   11: [NEQ(MV_MV12R.DriveBits,0) OTE(MV_MV12R.CW.[CWD.AUTODRV]) ,[XIC(MV_MV12R.CW.[CWD.AUTODRV]) XIO(MV_MV12R.CW.[CWD.MANUAL]) ,XIC(MV_MV12R.CW.[CWD.MANDRV]) XIC(MV_MV12R.CW.[CWD.MANUAL]) ] OTE(MV_MV12R.CW.[CWD.OUTPUT]) ,XIC(MV_MV12R.CW.[CWD.OUTPUT]) OTE(MV_MV12R_D) ,XIC(S:FS) [OTU(MV_MV12R.CW.[CWD.MANUAL]) ,LEQ(MV_MV12R.CheckTime,0) MOV(Default_Check_Time,MV_MV12R.CheckTime) ] ,[[XIC(MV_MV12R_R) XIO(Item_Simulation_Flag) ,XIC(Item_Simulation_Flag) [XIC(MV_MV12R.CW.[CWD.OUTPUT]) XIO(MV_MV12R.CW.[CWD.SIMFAIL]) ,XIO(MV_MV12R.CW.[CWD.OUTPUT]) XIC(MV_MV12R.CW.[CWD.SIMFAIL]) ] ] OTE(MV_MV12R.CW.[CWD.RUNFB]) ,[XIC(Item_Simulation_Flag) ,XIC(MV_MV12R.CW.[CWD.CHECKOFF]) ,XIC(Unused_Healthy_Feedback) ] OTE(MV_MV12R.CW.[CWD.HEALTHYFB]) ,[XIC(Item_Simulation_Flag) ,XIC(MV_MV12R.CW.[CWD.CHECKOFF]) ,XIC(Unused_NotTripped_Feedback) ] OTE(MV_MV12R.CW.[CWD.NOTTRIPPEDFB]) ] ,[XIC(MV_MV12R.CW.[CWD.AUTODRV]) XIO(MV_MV12R.CW.[CWD.PREVSCAN]) ,XIO(MV_MV12R.CW.[CWD.AUTODRV]) XIC(MV_MV12R.CW.[CWD.PREVSCAN]) ] CLR(MV_MV12R.CheckTimer) ,XIC(One_Second_One_Scan) LES(MV_MV12R.CheckTimer,MV_MV12R.CheckTime) ADD(MV_MV12R.CheckTimer,1,MV_MV12R.CheckTimer) ,XIO(MV_MV12R.CW.[CWD.FAULT]) OTU(MV_MV12R.CW.[CWD.FAULTLOGGED]) ,[GEQ(MV_MV12R.CheckTimer,MV_MV12R.CheckTime) [XIC(MV_MV12R.CW.[CWD.OUTPUT]) XIO(MV_MV12R.CW.[CWD.RUNFB]) ,XIO(MV_MV12R.CW.[CWD.OUTPUT]) XIC(MV_MV12R.CW.[CWD.RUNFB]) ] ,XIO(MV_MV12R.CW.[CWD.HEALTHYFB]) ,XIO(MV_MV12R.CW.[CWD.NOTTRIPPEDFB]) ,XIC(MV_MV12R.CW.[CWD.FAULT]) XIC(Item_Faults_Are_Latched) ,XIC(MV_MV12R.CW.[CWD.HIGHLIGHT]) ] XIO(MV_MV12R.CW.[CWD.CHECKOFF]) XIO(Alarm_Reset) [OTE(MV_MV12R.CW.[CWD.FAULT]) ,ALMD(MV_MV12R_ALARM,0,0,0,0) ] ,XIC(MV_MV12R.CW.[CWD.OUTPUT]) OTE(MV_MV12R.CW.[CWD.PREVSCAN]) ,XIC(MV_MV12R.CW.[CWD.FAULT]) EQU(Scada_Pump_Fault_No,0) XIO(MV_MV12R.CW.[CWD.FAULTLOGGED]) [MOV(20001,Scada_Pump_Fault_No) ,OTL(MV_MV12R.CW.[CWD.FAULTLOGGED]) ] ,XIO(MV_MV12R.CW.[CWD.HEALTHYFB]) EQU(Scada_Pump_H_Fault_No,0) XIO(MV_MV12R.CW.[CWD.HEALTHYFAULTLOGGED]) [MOV(20001,Scada_Pump_H_Fault_No) ,OTL(MV_MV12R.CW.[CWD.HEALTHYFAULTLOGGED]) ] ,XIO(MV_MV12R.CW.[CWD.NOTTRIPPEDFB]) EQU(Scada_Pump_H_Fault_No,0) XIO(MV_MV12R.CW.[CWD.TRIPPEDFAULTLOGGED]) [MOV(20001,Scada_Pump_T_Fault_No) ,OTL(MV_MV12R.CW.[CWD.TRIPPEDFAULTLOGGED]) ] ];
   12: [NEQ(MV_MV13R.DriveBits,0) OTE(MV_MV13R.CW.[CWD.AUTODRV]) ,[XIC(MV_MV13R.CW.[CWD.AUTODRV]) XIO(MV_MV13R.CW.[CWD.MANUAL]) ,XIC(MV_MV13R.CW.[CWD.MANDRV]) XIC(MV_MV13R.CW.[CWD.MANUAL]) ] OTE(MV_MV13R.CW.[CWD.OUTPUT]) ,XIC(MV_MV13R.CW.[CWD.OUTPUT]) OTE(MV_MV13R_D) ,XIC(S:FS) [OTU(MV_MV13R.CW.[CWD.MANUAL]) ,LEQ(MV_MV13R.CheckTime,0) MOV(Default_Check_Time,MV_MV13R.CheckTime) ] ,[[XIC(MV_MV13R_R) XIO(Item_Simulation_Flag) ,XIC(Item_Simulation_Flag) [XIC(MV_MV13R.CW.[CWD.OUTPUT]) XIO(MV_MV13R.CW.[CWD.SIMFAIL]) ,XIO(MV_MV13R.CW.[CWD.OUTPUT]) XIC(MV_MV13R.CW.[CWD.SIMFAIL]) ] ] OTE(MV_MV13R.CW.[CWD.RUNFB]) ,[XIC(Item_Simulation_Flag) ,XIC(MV_MV13R.CW.[CWD.CHECKOFF]) ,XIC(Unused_Healthy_Feedback) ] OTE(MV_MV13R.CW.[CWD.HEALTHYFB]) ,[XIC(Item_Simulation_Flag) ,XIC(MV_MV13R.CW.[CWD.CHECKOFF]) ,XIC(Unused_NotTripped_Feedback) ] OTE(MV_MV13R.CW.[CWD.NOTTRIPPEDFB]) ] ,[XIC(MV_MV13R.CW.[CWD.AUTODRV]) XIO(MV_MV13R.CW.[CWD.PREVSCAN]) ,XIO(MV_MV13R.CW.[CWD.AUTODRV]) XIC(MV_MV13R.CW.[CWD.PREVSCAN]) ] CLR(MV_MV13R.CheckTimer) ,XIC(One_Second_One_Scan) LES(MV_MV13R.CheckTimer,MV_MV13R.CheckTime) ADD(MV_MV13R.CheckTimer,1,MV_MV13R.CheckTimer) ,XIO(MV_MV13R.CW.[CWD.FAULT]) OTU(MV_MV13R.CW.[CWD.FAULTLOGGED]) ,[GEQ(MV_MV13R.CheckTimer,MV_MV13R.CheckTime) [XIC(MV_MV13R.CW.[CWD.OUTPUT]) XIO(MV_MV13R.CW.[CWD.RUNFB]) ,XIO(MV_MV13R.CW.[CWD.OUTPUT]) XIC(MV_MV13R.CW.[CWD.RUNFB]) ] ,XIO(MV_MV13R.CW.[CWD.HEALTHYFB]) ,XIO(MV_MV13R.CW.[CWD.NOTTRIPPEDFB]) ,XIC(MV_MV13R.CW.[CWD.FAULT]) XIC(Item_Faults_Are_Latched) ,XIC(MV_MV13R.CW.[CWD.HIGHLIGHT]) ] XIO(MV_MV13R.CW.[CWD.CHECKOFF]) XIO(Alarm_Reset) [OTE(MV_MV13R.CW.[CWD.FAULT]) ,ALMD(MV_MV13R_ALARM,0,0,0,0) ] ,XIC(MV_MV13R.CW.[CWD.OUTPUT]) OTE(MV_MV13R.CW.[CWD.PREVSCAN]) ,XIC(MV_MV13R.CW.[CWD.FAULT]) EQU(Scada_Pump_Fault_No,0) XIO(MV_MV13R.CW.[CWD.FAULTLOGGED]) [MOV(20001,Scada_Pump_Fault_No) ,OTL(MV_MV13R.CW.[CWD.FAULTLOGGED]) ] ,XIO(MV_MV13R.CW.[CWD.HEALTHYFB]) EQU(Scada_Pump_H_Fault_No,0) XIO(MV_MV13R.CW.[CWD.HEALTHYFAULTLOGGED]) [MOV(20001,Scada_Pump_H_Fault_No) ,OTL(MV_MV13R.CW.[CWD.HEALTHYFAULTLOGGED]) ] ,XIO(MV_MV13R.CW.[CWD.NOTTRIPPEDFB]) EQU(Scada_Pump_H_Fault_No,0) XIO(MV_MV13R.CW.[CWD.TRIPPEDFAULTLOGGED]) [MOV(20001,Scada_Pump_T_Fault_No) ,OTL(MV_MV13R.CW.[CWD.TRIPPEDFAULTLOGGED]) ] ];
   13: [NEQ(MV_MV14R.DriveBits,0) OTE(MV_MV14R.CW.[CWD.AUTODRV]) ,[XIC(MV_MV14R.CW.[CWD.AUTODRV]) XIO(MV_MV14R.CW.[CWD.MANUAL]) ,XIC(MV_MV14R.CW.[CWD.MANDRV]) XIC(MV_MV14R.CW.[CWD.MANUAL]) ] OTE(MV_MV14R.CW.[CWD.OUTPUT]) ,XIC(MV_MV14R.CW.[CWD.OUTPUT]) OTE(MV_MV14R_D) ,XIC(S:FS) [OTU(MV_MV14R.CW.[CWD.MANUAL]) ,LEQ(MV_MV14R.CheckTime,0) MOV(Default_Check_Time,MV_MV14R.CheckTime) ] ,[[XIC(MV_MV14R_R) XIO(Item_Simulation_Flag) ,XIC(Item_Simulation_Flag) [XIC(MV_MV14R.CW.[CWD.OUTPUT]) XIO(MV_MV14R.CW.[CWD.SIMFAIL]) ,XIO(MV_MV14R.CW.[CWD.OUTPUT]) XIC(MV_MV14R.CW.[CWD.SIMFAIL]) ] ] OTE(MV_MV14R.CW.[CWD.RUNFB]) ,[XIC(Item_Simulation_Flag) ,XIC(MV_MV14R.CW.[CWD.CHECKOFF]) ,XIC(Unused_Healthy_Feedback) ] OTE(MV_MV14R.CW.[CWD.HEALTHYFB]) ,[XIC(Item_Simulation_Flag) ,XIC(MV_MV14R.CW.[CWD.CHECKOFF]) ,XIC(Unused_NotTripped_Feedback) ] OTE(MV_MV14R.CW.[CWD.NOTTRIPPEDFB]) ] ,[XIC(MV_MV14R.CW.[CWD.AUTODRV]) XIO(MV_MV14R.CW.[CWD.PREVSCAN]) ,XIO(MV_MV14R.CW.[CWD.AUTODRV]) XIC(MV_MV14R.CW.[CWD.PREVSCAN]) ] CLR(MV_MV14R.CheckTimer) ,XIC(One_Second_One_Scan) LES(MV_MV14R.CheckTimer,MV_MV14R.CheckTime) ADD(MV_MV14R.CheckTimer,1,MV_MV14R.CheckTimer) ,XIO(MV_MV14R.CW.[CWD.FAULT]) OTU(MV_MV14R.CW.[CWD.FAULTLOGGED]) ,[GEQ(MV_MV14R.CheckTimer,MV_MV14R.CheckTime) [XIC(MV_MV14R.CW.[CWD.OUTPUT]) XIO(MV_MV14R.CW.[CWD.RUNFB]) ,XIO(MV_MV14R.CW.[CWD.OUTPUT]) XIC(MV_MV14R.CW.[CWD.RUNFB]) ] ,XIO(MV_MV14R.CW.[CWD.HEALTHYFB]) ,XIO(MV_MV14R.CW.[CWD.NOTTRIPPEDFB]) ,XIC(MV_MV14R.CW.[CWD.FAULT]) XIC(Item_Faults_Are_Latched) ,XIC(MV_MV14R.CW.[CWD.HIGHLIGHT]) ] XIO(MV_MV14R.CW.[CWD.CHECKOFF]) XIO(Alarm_Reset) [OTE(MV_MV14R.CW.[CWD.FAULT]) ,ALMD(MV_MV14R_ALARM,0,0,0,0) ] ,XIC(MV_MV14R.CW.[CWD.OUTPUT]) OTE(MV_MV14R.CW.[CWD.PREVSCAN]) ,XIC(MV_MV14R.CW.[CWD.FAULT]) EQU(Scada_Pump_Fault_No,0) XIO(MV_MV14R.CW.[CWD.FAULTLOGGED]) [MOV(20001,Scada_Pump_Fault_No) ,OTL(MV_MV14R.CW.[CWD.FAULTLOGGED]) ] ,XIO(MV_MV14R.CW.[CWD.HEALTHYFB]) EQU(Scada_Pump_H_Fault_No,0) XIO(MV_MV14R.CW.[CWD.HEALTHYFAULTLOGGED]) [MOV(20001,Scada_Pump_H_Fault_No) ,OTL(MV_MV14R.CW.[CWD.HEALTHYFAULTLOGGED]) ] ,XIO(MV_MV14R.CW.[CWD.NOTTRIPPEDFB]) EQU(Scada_Pump_H_Fault_No,0) XIO(MV_MV14R.CW.[CWD.TRIPPEDFAULTLOGGED]) [MOV(20001,Scada_Pump_T_Fault_No) ,OTL(MV_MV14R.CW.[CWD.TRIPPEDFAULTLOGGED]) ] ];
   14: [NEQ(MV_MV15R.DriveBits,0) OTE(MV_MV15R.CW.[CWD.AUTODRV]) ,[XIC(MV_MV15R.CW.[CWD.AUTODRV]) XIO(MV_MV15R.CW.[CWD.MANUAL]) ,XIC(MV_MV15R.CW.[CWD.MANDRV]) XIC(MV_MV15R.CW.[CWD.MANUAL]) ] OTE(MV_MV15R.CW.[CWD.OUTPUT]) ,XIC(MV_MV15R.CW.[CWD.OUTPUT]) OTE(MV_MV15R_D) ,XIC(S:FS) [OTU(MV_MV15R.CW.[CWD.MANUAL]) ,LEQ(MV_MV15R.CheckTime,0) MOV(Default_Check_Time,MV_MV15R.CheckTime) ] ,[[XIC(MV_MV15R_R) XIO(Item_Simulation_Flag) ,XIC(Item_Simulation_Flag) [XIC(MV_MV15R.CW.[CWD.OUTPUT]) XIO(MV_MV15R.CW.[CWD.SIMFAIL]) ,XIO(MV_MV15R.CW.[CWD.OUTPUT]) XIC(MV_MV15R.CW.[CWD.SIMFAIL]) ] ] OTE(MV_MV15R.CW.[CWD.RUNFB]) ,[XIC(Item_Simulation_Flag) ,XIC(MV_MV15R.CW.[CWD.CHECKOFF]) ,XIC(Unused_Healthy_Feedback) ] OTE(MV_MV15R.CW.[CWD.HEALTHYFB]) ,[XIC(Item_Simulation_Flag) ,XIC(MV_MV15R.CW.[CWD.CHECKOFF]) ,XIC(Unused_NotTripped_Feedback) ] OTE(MV_MV15R.CW.[CWD.NOTTRIPPEDFB]) ] ,[XIC(MV_MV15R.CW.[CWD.AUTODRV]) XIO(MV_MV15R.CW.[CWD.PREVSCAN]) ,XIO(MV_MV15R.CW.[CWD.AUTODRV]) XIC(MV_MV15R.CW.[CWD.PREVSCAN]) ] CLR(MV_MV15R.CheckTimer) ,XIC(One_Second_One_Scan) LES(MV_MV15R.CheckTimer,MV_MV15R.CheckTime) ADD(MV_MV15R.CheckTimer,1,MV_MV15R.CheckTimer) ,XIO(MV_MV15R.CW.[CWD.FAULT]) OTU(MV_MV15R.CW.[CWD.FAULTLOGGED]) ,[GEQ(MV_MV15R.CheckTimer,MV_MV15R.CheckTime) [XIC(MV_MV15R.CW.[CWD.OUTPUT]) XIO(MV_MV15R.CW.[CWD.RUNFB]) ,XIO(MV_MV15R.CW.[CWD.OUTPUT]) XIC(MV_MV15R.CW.[CWD.RUNFB]) ] ,XIO(MV_MV15R.CW.[CWD.HEALTHYFB]) ,XIO(MV_MV15R.CW.[CWD.NOTTRIPPEDFB]) ,XIC(MV_MV15R.CW.[CWD.FAULT]) XIC(Item_Faults_Are_Latched) ,XIC(MV_MV15R.CW.[CWD.HIGHLIGHT]) ] XIO(MV_MV15R.CW.[CWD.CHECKOFF]) XIO(Alarm_Reset) [OTE(MV_MV15R.CW.[CWD.FAULT]) ,ALMD(MV_MV15R_ALARM,0,0,0,0) ] ,XIC(MV_MV15R.CW.[CWD.OUTPUT]) OTE(MV_MV15R.CW.[CWD.PREVSCAN]) ,XIC(MV_MV15R.CW.[CWD.FAULT]) EQU(Scada_Pump_Fault_No,0) XIO(MV_MV15R.CW.[CWD.FAULTLOGGED]) [MOV(20001,Scada_Pump_Fault_No) ,OTL(MV_MV15R.CW.[CWD.FAULTLOGGED]) ] ,XIO(MV_MV15R.CW.[CWD.HEALTHYFB]) EQU(Scada_Pump_H_Fault_No,0) XIO(MV_MV15R.CW.[CWD.HEALTHYFAULTLOGGED]) [MOV(20001,Scada_Pump_H_Fault_No) ,OTL(MV_MV15R.CW.[CWD.HEALTHYFAULTLOGGED]) ] ,XIO(MV_MV15R.CW.[CWD.NOTTRIPPEDFB]) EQU(Scada_Pump_H_Fault_No,0) XIO(MV_MV15R.CW.[CWD.TRIPPEDFAULTLOGGED]) [MOV(20001,Scada_Pump_T_Fault_No) ,OTL(MV_MV15R.CW.[CWD.TRIPPEDFAULTLOGGED]) ] ];
   15: [NEQ(MV_MV16R.DriveBits,0) OTE(MV_MV16R.CW.[CWD.AUTODRV]) ,[XIC(MV_MV16R.CW.[CWD.AUTODRV]) XIO(MV_MV16R.CW.[CWD.MANUAL]) ,XIC(MV_MV16R.CW.[CWD.MANDRV]) XIC(MV_MV16R.CW.[CWD.MANUAL]) ] OTE(MV_MV16R.CW.[CWD.OUTPUT]) ,XIC(MV_MV16R.CW.[CWD.OUTPUT]) OTE(MV_MV16R_D) ,XIC(S:FS) [OTU(MV_MV16R.CW.[CWD.MANUAL]) ,LEQ(MV_MV16R.CheckTime,0) MOV(Default_Check_Time,MV_MV16R.CheckTime) ] ,[[XIC(MV_MV16R_R) XIO(Item_Simulation_Flag) ,XIC(Item_Simulation_Flag) [XIC(MV_MV16R.CW.[CWD.OUTPUT]) XIO(MV_MV16R.CW.[CWD.SIMFAIL]) ,XIO(MV_MV16R.CW.[CWD.OUTPUT]) XIC(MV_MV16R.CW.[CWD.SIMFAIL]) ] ] OTE(MV_MV16R.CW.[CWD.RUNFB]) ,[XIC(Item_Simulation_Flag) ,XIC(MV_MV16R.CW.[CWD.CHECKOFF]) ,XIC(Unused_Healthy_Feedback) ] OTE(MV_MV16R.CW.[CWD.HEALTHYFB]) ,[XIC(Item_Simulation_Flag) ,XIC(MV_MV16R.CW.[CWD.CHECKOFF]) ,XIC(Unused_NotTripped_Feedback) ] OTE(MV_MV16R.CW.[CWD.NOTTRIPPEDFB]) ] ,[XIC(MV_MV16R.CW.[CWD.AUTODRV]) XIO(MV_MV16R.CW.[CWD.PREVSCAN]) ,XIO(MV_MV16R.CW.[CWD.AUTODRV]) XIC(MV_MV16R.CW.[CWD.PREVSCAN]) ] CLR(MV_MV16R.CheckTimer) ,XIC(One_Second_One_Scan) LES(MV_MV16R.CheckTimer,MV_MV16R.CheckTime) ADD(MV_MV16R.CheckTimer,1,MV_MV16R.CheckTimer) ,XIO(MV_MV16R.CW.[CWD.FAULT]) OTU(MV_MV16R.CW.[CWD.FAULTLOGGED]) ,[GEQ(MV_MV16R.CheckTimer,MV_MV16R.CheckTime) [XIC(MV_MV16R.CW.[CWD.OUTPUT]) XIO(MV_MV16R.CW.[CWD.RUNFB]) ,XIO(MV_MV16R.CW.[CWD.OUTPUT]) XIC(MV_MV16R.CW.[CWD.RUNFB]) ] ,XIO(MV_MV16R.CW.[CWD.HEALTHYFB]) ,XIO(MV_MV16R.CW.[CWD.NOTTRIPPEDFB]) ,XIC(MV_MV16R.CW.[CWD.FAULT]) XIC(Item_Faults_Are_Latched) ,XIC(MV_MV16R.CW.[CWD.HIGHLIGHT]) ] XIO(MV_MV16R.CW.[CWD.CHECKOFF]) XIO(Alarm_Reset) [OTE(MV_MV16R.CW.[CWD.FAULT]) ,ALMD(MV_MV16R_ALARM,0,0,0,0) ] ,XIC(MV_MV16R.CW.[CWD.OUTPUT]) OTE(MV_MV16R.CW.[CWD.PREVSCAN]) ,XIC(MV_MV16R.CW.[CWD.FAULT]) EQU(Scada_Pump_Fault_No,0) XIO(MV_MV16R.CW.[CWD.FAULTLOGGED]) [MOV(20001,Scada_Pump_Fault_No) ,OTL(MV_MV16R.CW.[CWD.FAULTLOGGED]) ] ,XIO(MV_MV16R.CW.[CWD.HEALTHYFB]) EQU(Scada_Pump_H_Fault_No,0) XIO(MV_MV16R.CW.[CWD.HEALTHYFAULTLOGGED]) [MOV(20001,Scada_Pump_H_Fault_No) ,OTL(MV_MV16R.CW.[CWD.HEALTHYFAULTLOGGED]) ] ,XIO(MV_MV16R.CW.[CWD.NOTTRIPPEDFB]) EQU(Scada_Pump_H_Fault_No,0) XIO(MV_MV16R.CW.[CWD.TRIPPEDFAULTLOGGED]) [MOV(20001,Scada_Pump_T_Fault_No) ,OTL(MV_MV16R.CW.[CWD.TRIPPEDFAULTLOGGED]) ] ];
   16: [NEQ(MV_MV17R.DriveBits,0) OTE(MV_MV17R.CW.[CWD.AUTODRV]) ,[XIC(MV_MV17R.CW.[CWD.AUTODRV]) XIO(MV_MV17R.CW.[CWD.MANUAL]) ,XIC(MV_MV17R.CW.[CWD.MANDRV]) XIC(MV_MV17R.CW.[CWD.MANUAL]) ] OTE(MV_MV17R.CW.[CWD.OUTPUT]) ,XIC(MV_MV17R.CW.[CWD.OUTPUT]) OTE(MV_MV17R_D) ,XIC(S:FS) [OTU(MV_MV17R.CW.[CWD.MANUAL]) ,LEQ(MV_MV17R.CheckTime,0) MOV(Default_Check_Time,MV_MV17R.CheckTime) ] ,[[XIC(MV_MV17R_R) XIO(Item_Simulation_Flag) ,XIC(Item_Simulation_Flag) [XIC(MV_MV17R.CW.[CWD.OUTPUT]) XIO(MV_MV17R.CW.[CWD.SIMFAIL]) ,XIO(MV_MV17R.CW.[CWD.OUTPUT]) XIC(MV_MV17R.CW.[CWD.SIMFAIL]) ] ] OTE(MV_MV17R.CW.[CWD.RUNFB]) ,[XIC(Item_Simulation_Flag) ,XIC(MV_MV17R.CW.[CWD.CHECKOFF]) ,XIC(Unused_Healthy_Feedback) ] OTE(MV_MV17R.CW.[CWD.HEALTHYFB]) ,[XIC(Item_Simulation_Flag) ,XIC(MV_MV17R.CW.[CWD.CHECKOFF]) ,XIC(Unused_NotTripped_Feedback) ] OTE(MV_MV17R.CW.[CWD.NOTTRIPPEDFB]) ] ,[XIC(MV_MV17R.CW.[CWD.AUTODRV]) XIO(MV_MV17R.CW.[CWD.PREVSCAN]) ,XIO(MV_MV17R.CW.[CWD.AUTODRV]) XIC(MV_MV17R.CW.[CWD.PREVSCAN]) ] CLR(MV_MV17R.CheckTimer) ,XIC(One_Second_One_Scan) LES(MV_MV17R.CheckTimer,MV_MV17R.CheckTime) ADD(MV_MV17R.CheckTimer,1,MV_MV17R.CheckTimer) ,XIO(MV_MV17R.CW.[CWD.FAULT]) OTU(MV_MV17R.CW.[CWD.FAULTLOGGED]) ,[GEQ(MV_MV17R.CheckTimer,MV_MV17R.CheckTime) [XIC(MV_MV17R.CW.[CWD.OUTPUT]) XIO(MV_MV17R.CW.[CWD.RUNFB]) ,XIO(MV_MV17R.CW.[CWD.OUTPUT]) XIC(MV_MV17R.CW.[CWD.RUNFB]) ] ,XIO(MV_MV17R.CW.[CWD.HEALTHYFB]) ,XIO(MV_MV17R.CW.[CWD.NOTTRIPPEDFB]) ,XIC(MV_MV17R.CW.[CWD.FAULT]) XIC(Item_Faults_Are_Latched) ,XIC(MV_MV17R.CW.[CWD.HIGHLIGHT]) ] XIO(MV_MV17R.CW.[CWD.CHECKOFF]) XIO(Alarm_Reset) [OTE(MV_MV17R.CW.[CWD.FAULT]) ,ALMD(MV_MV17R_ALARM,0,0,0,0) ] ,XIC(MV_MV17R.CW.[CWD.OUTPUT]) OTE(MV_MV17R.CW.[CWD.PREVSCAN]) ,XIC(MV_MV17R.CW.[CWD.FAULT]) EQU(Scada_Pump_Fault_No,0) XIO(MV_MV17R.CW.[CWD.FAULTLOGGED]) [MOV(20001,Scada_Pump_Fault_No) ,OTL(MV_MV17R.CW.[CWD.FAULTLOGGED]) ] ,XIO(MV_MV17R.CW.[CWD.HEALTHYFB]) EQU(Scada_Pump_H_Fault_No,0) XIO(MV_MV17R.CW.[CWD.HEALTHYFAULTLOGGED]) [MOV(20001,Scada_Pump_H_Fault_No) ,OTL(MV_MV17R.CW.[CWD.HEALTHYFAULTLOGGED]) ] ,XIO(MV_MV17R.CW.[CWD.NOTTRIPPEDFB]) EQU(Scada_Pump_H_Fault_No,0) XIO(MV_MV17R.CW.[CWD.TRIPPEDFAULTLOGGED]) [MOV(20001,Scada_Pump_T_Fault_No) ,OTL(MV_MV17R.CW.[CWD.TRIPPEDFAULTLOGGED]) ] ];
   17: [NEQ(MV_MV18R.DriveBits,0) OTE(MV_MV18R.CW.[CWD.AUTODRV]) ,[XIC(MV_MV18R.CW.[CWD.AUTODRV]) XIO(MV_MV18R.CW.[CWD.MANUAL]) ,XIC(MV_MV18R.CW.[CWD.MANDRV]) XIC(MV_MV18R.CW.[CWD.MANUAL]) ] OTE(MV_MV18R.CW.[CWD.OUTPUT]) ,XIC(MV_MV18R.CW.[CWD.OUTPUT]) OTE(MV_MV18R_D) ,XIC(S:FS) [OTU(MV_MV18R.CW.[CWD.MANUAL]) ,LEQ(MV_MV18R.CheckTime,0) MOV(Default_Check_Time,MV_MV18R.CheckTime) ] ,[[XIC(MV_MV18R_R) XIO(Item_Simulation_Flag) ,XIC(Item_Simulation_Flag) [XIC(MV_MV18R.CW.[CWD.OUTPUT]) XIO(MV_MV18R.CW.[CWD.SIMFAIL]) ,XIO(MV_MV18R.CW.[CWD.OUTPUT]) XIC(MV_MV18R.CW.[CWD.SIMFAIL]) ] ] OTE(MV_MV18R.CW.[CWD.RUNFB]) ,[XIC(Item_Simulation_Flag) ,XIC(MV_MV18R.CW.[CWD.CHECKOFF]) ,XIC(Unused_Healthy_Feedback) ] OTE(MV_MV18R.CW.[CWD.HEALTHYFB]) ,[XIC(Item_Simulation_Flag) ,XIC(MV_MV18R.CW.[CWD.CHECKOFF]) ,XIC(Unused_NotTripped_Feedback) ] OTE(MV_MV18R.CW.[CWD.NOTTRIPPEDFB]) ] ,[XIC(MV_MV18R.CW.[CWD.AUTODRV]) XIO(MV_MV18R.CW.[CWD.PREVSCAN]) ,XIO(MV_MV18R.CW.[CWD.AUTODRV]) XIC(MV_MV18R.CW.[CWD.PREVSCAN]) ] CLR(MV_MV18R.CheckTimer) ,XIC(One_Second_One_Scan) LES(MV_MV18R.CheckTimer,MV_MV18R.CheckTime) ADD(MV_MV18R.CheckTimer,1,MV_MV18R.CheckTimer) ,XIO(MV_MV18R.CW.[CWD.FAULT]) OTU(MV_MV18R.CW.[CWD.FAULTLOGGED]) ,[GEQ(MV_MV18R.CheckTimer,MV_MV18R.CheckTime) [XIC(MV_MV18R.CW.[CWD.OUTPUT]) XIO(MV_MV18R.CW.[CWD.RUNFB]) ,XIO(MV_MV18R.CW.[CWD.OUTPUT]) XIC(MV_MV18R.CW.[CWD.RUNFB]) ] ,XIO(MV_MV18R.CW.[CWD.HEALTHYFB]) ,XIO(MV_MV18R.CW.[CWD.NOTTRIPPEDFB]) ,XIC(MV_MV18R.CW.[CWD.FAULT]) XIC(Item_Faults_Are_Latched) ,XIC(MV_MV18R.CW.[CWD.HIGHLIGHT]) ] XIO(MV_MV18R.CW.[CWD.CHECKOFF]) XIO(Alarm_Reset) [OTE(MV_MV18R.CW.[CWD.FAULT]) ,ALMD(MV_MV18R_ALARM,0,0,0,0) ] ,XIC(MV_MV18R.CW.[CWD.OUTPUT]) OTE(MV_MV18R.CW.[CWD.PREVSCAN]) ,XIC(MV_MV18R.CW.[CWD.FAULT]) EQU(Scada_Pump_Fault_No,0) XIO(MV_MV18R.CW.[CWD.FAULTLOGGED]) [MOV(20001,Scada_Pump_Fault_No) ,OTL(MV_MV18R.CW.[CWD.FAULTLOGGED]) ] ,XIO(MV_MV18R.CW.[CWD.HEALTHYFB]) EQU(Scada_Pump_H_Fault_No,0) XIO(MV_MV18R.CW.[CWD.HEALTHYFAULTLOGGED]) [MOV(20001,Scada_Pump_H_Fault_No) ,OTL(MV_MV18R.CW.[CWD.HEALTHYFAULTLOGGED]) ] ,XIO(MV_MV18R.CW.[CWD.NOTTRIPPEDFB]) EQU(Scada_Pump_H_Fault_No,0) XIO(MV_MV18R.CW.[CWD.TRIPPEDFAULTLOGGED]) [MOV(20001,Scada_Pump_T_Fault_No) ,OTL(MV_MV18R.CW.[CWD.TRIPPEDFAULTLOGGED]) ] ];
   18: [NEQ(MV_MV19R.DriveBits,0) OTE(MV_MV19R.CW.[CWD.AUTODRV]) ,[XIC(MV_MV19R.CW.[CWD.AUTODRV]) XIO(MV_MV19R.CW.[CWD.MANUAL]) ,XIC(MV_MV19R.CW.[CWD.MANDRV]) XIC(MV_MV19R.CW.[CWD.MANUAL]) ] OTE(MV_MV19R.CW.[CWD.OUTPUT]) ,XIC(MV_MV19R.CW.[CWD.OUTPUT]) OTE(MV_MV19R_D) ,XIC(S:FS) [OTU(MV_MV19R.CW.[CWD.MANUAL]) ,LEQ(MV_MV19R.CheckTime,0) MOV(Default_Check_Time,MV_MV19R.CheckTime) ] ,[[XIC(MV_MV19R_R) XIO(Item_Simulation_Flag) ,XIC(Item_Simulation_Flag) [XIC(MV_MV19R.CW.[CWD.OUTPUT]) XIO(MV_MV19R.CW.[CWD.SIMFAIL]) ,XIO(MV_MV19R.CW.[CWD.OUTPUT]) XIC(MV_MV19R.CW.[CWD.SIMFAIL]) ] ] OTE(MV_MV19R.CW.[CWD.RUNFB]) ,[XIC(Item_Simulation_Flag) ,XIC(MV_MV19R.CW.[CWD.CHECKOFF]) ,XIC(Unused_Healthy_Feedback) ] OTE(MV_MV19R.CW.[CWD.HEALTHYFB]) ,[XIC(Item_Simulation_Flag) ,XIC(MV_MV19R.CW.[CWD.CHECKOFF]) ,XIC(Unused_NotTripped_Feedback) ] OTE(MV_MV19R.CW.[CWD.NOTTRIPPEDFB]) ] ,[XIC(MV_MV19R.CW.[CWD.AUTODRV]) XIO(MV_MV19R.CW.[CWD.PREVSCAN]) ,XIO(MV_MV19R.CW.[CWD.AUTODRV]) XIC(MV_MV19R.CW.[CWD.PREVSCAN]) ] CLR(MV_MV19R.CheckTimer) ,XIC(One_Second_One_Scan) LES(MV_MV19R.CheckTimer,MV_MV19R.CheckTime) ADD(MV_MV19R.CheckTimer,1,MV_MV19R.CheckTimer) ,XIO(MV_MV19R.CW.[CWD.FAULT]) OTU(MV_MV19R.CW.[CWD.FAULTLOGGED]) ,[GEQ(MV_MV19R.CheckTimer,MV_MV19R.CheckTime) [XIC(MV_MV19R.CW.[CWD.OUTPUT]) XIO(MV_MV19R.CW.[CWD.RUNFB]) ,XIO(MV_MV19R.CW.[CWD.OUTPUT]) XIC(MV_MV19R.CW.[CWD.RUNFB]) ] ,XIO(MV_MV19R.CW.[CWD.HEALTHYFB]) ,XIO(MV_MV19R.CW.[CWD.NOTTRIPPEDFB]) ,XIC(MV_MV19R.CW.[CWD.FAULT]) XIC(Item_Faults_Are_Latched) ,XIC(MV_MV19R.CW.[CWD.HIGHLIGHT]) ] XIO(MV_MV19R.CW.[CWD.CHECKOFF]) XIO(Alarm_Reset) [OTE(MV_MV19R.CW.[CWD.FAULT]) ,ALMD(MV_MV19R_ALARM,0,0,0,0) ] ,XIC(MV_MV19R.CW.[CWD.OUTPUT]) OTE(MV_MV19R.CW.[CWD.PREVSCAN]) ,XIC(MV_MV19R.CW.[CWD.FAULT]) EQU(Scada_Pump_Fault_No,0) XIO(MV_MV19R.CW.[CWD.FAULTLOGGED]) [MOV(20001,Scada_Pump_Fault_No) ,OTL(MV_MV19R.CW.[CWD.FAULTLOGGED]) ] ,XIO(MV_MV19R.CW.[CWD.HEALTHYFB]) EQU(Scada_Pump_H_Fault_No,0) XIO(MV_MV19R.CW.[CWD.HEALTHYFAULTLOGGED]) [MOV(20001,Scada_Pump_H_Fault_No) ,OTL(MV_MV19R.CW.[CWD.HEALTHYFAULTLOGGED]) ] ,XIO(MV_MV19R.CW.[CWD.NOTTRIPPEDFB]) EQU(Scada_Pump_H_Fault_No,0) XIO(MV_MV19R.CW.[CWD.TRIPPEDFAULTLOGGED]) [MOV(20001,Scada_Pump_T_Fault_No) ,OTL(MV_MV19R.CW.[CWD.TRIPPEDFAULTLOGGED]) ] ];
   19: [NEQ(MV_MV30R.DriveBits,0) OTE(MV_MV30R.CW.[CWD.AUTODRV]) ,[XIC(MV_MV30R.CW.[CWD.AUTODRV]) XIO(MV_MV30R.CW.[CWD.MANUAL]) ,XIC(MV_MV30R.CW.[CWD.MANDRV]) XIC(MV_MV30R.CW.[CWD.MANUAL]) ] OTE(MV_MV30R.CW.[CWD.OUTPUT]) ,XIC(MV_MV30R.CW.[CWD.OUTPUT]) OTE(MV_MV30R_D) ,XIC(S:FS) [OTU(MV_MV30R.CW.[CWD.MANUAL]) ,LEQ(MV_MV30R.CheckTime,0) MOV(Default_Check_Time,MV_MV30R.CheckTime) ] ,[[XIC(MV_MV30R_R) XIO(Item_Simulation_Flag) ,XIC(Item_Simulation_Flag) [XIC(MV_MV30R.CW.[CWD.OUTPUT]) XIO(MV_MV30R.CW.[CWD.SIMFAIL]) ,XIO(MV_MV30R.CW.[CWD.OUTPUT]) XIC(MV_MV30R.CW.[CWD.SIMFAIL]) ] ] OTE(MV_MV30R.CW.[CWD.RUNFB]) ,[XIC(Item_Simulation_Flag) ,XIC(MV_MV30R.CW.[CWD.CHECKOFF]) ,XIC(Unused_Healthy_Feedback) ] OTE(MV_MV30R.CW.[CWD.HEALTHYFB]) ,[XIC(Item_Simulation_Flag) ,XIC(MV_MV30R.CW.[CWD.CHECKOFF]) ,XIC(Unused_NotTripped_Feedback) ] OTE(MV_MV30R.CW.[CWD.NOTTRIPPEDFB]) ] ,[XIC(MV_MV30R.CW.[CWD.AUTODRV]) XIO(MV_MV30R.CW.[CWD.PREVSCAN]) ,XIO(MV_MV30R.CW.[CWD.AUTODRV]) XIC(MV_MV30R.CW.[CWD.PREVSCAN]) ] CLR(MV_MV30R.CheckTimer) ,XIC(One_Second_One_Scan) LES(MV_MV30R.CheckTimer,MV_MV30R.CheckTime) ADD(MV_MV30R.CheckTimer,1,MV_MV30R.CheckTimer) ,XIO(MV_MV30R.CW.[CWD.FAULT]) OTU(MV_MV30R.CW.[CWD.FAULTLOGGED]) ,[GEQ(MV_MV30R.CheckTimer,MV_MV30R.CheckTime) [XIC(MV_MV30R.CW.[CWD.OUTPUT]) XIO(MV_MV30R.CW.[CWD.RUNFB]) ,XIO(MV_MV30R.CW.[CWD.OUTPUT]) XIC(MV_MV30R.CW.[CWD.RUNFB]) ] ,XIO(MV_MV30R.CW.[CWD.HEALTHYFB]) ,XIO(MV_MV30R.CW.[CWD.NOTTRIPPEDFB]) ,XIC(MV_MV30R.CW.[CWD.FAULT]) XIC(Item_Faults_Are_Latched) ,XIC(MV_MV30R.CW.[CWD.HIGHLIGHT]) ] XIO(MV_MV30R.CW.[CWD.CHECKOFF]) XIO(Alarm_Reset) [OTE(MV_MV30R.CW.[CWD.FAULT]) ,ALMD(MV_MV30R_ALARM,0,0,0,0) ] ,XIC(MV_MV30R.CW.[CWD.OUTPUT]) OTE(MV_MV30R.CW.[CWD.PREVSCAN]) ,XIC(MV_MV30R.CW.[CWD.FAULT]) EQU(Scada_Pump_Fault_No,0) XIO(MV_MV30R.CW.[CWD.FAULTLOGGED]) [MOV(20001,Scada_Pump_Fault_No) ,OTL(MV_MV30R.CW.[CWD.FAULTLOGGED]) ] ,XIO(MV_MV30R.CW.[CWD.HEALTHYFB]) EQU(Scada_Pump_H_Fault_No,0) XIO(MV_MV30R.CW.[CWD.HEALTHYFAULTLOGGED]) [MOV(20001,Scada_Pump_H_Fault_No) ,OTL(MV_MV30R.CW.[CWD.HEALTHYFAULTLOGGED]) ] ,XIO(MV_MV30R.CW.[CWD.NOTTRIPPEDFB]) EQU(Scada_Pump_H_Fault_No,0) XIO(MV_MV30R.CW.[CWD.TRIPPEDFAULTLOGGED]) [MOV(20001,Scada_Pump_T_Fault_No) ,OTL(MV_MV30R.CW.[CWD.TRIPPEDFAULTLOGGED]) ] ];
   20: [NEQ(MV_MV31R.DriveBits,0) OTE(MV_MV31R.CW.[CWD.AUTODRV]) ,[XIC(MV_MV31R.CW.[CWD.AUTODRV]) XIO(MV_MV31R.CW.[CWD.MANUAL]) ,XIC(MV_MV31R.CW.[CWD.MANDRV]) XIC(MV_MV31R.CW.[CWD.MANUAL]) ] OTE(MV_MV31R.CW.[CWD.OUTPUT]) ,XIC(MV_MV31R.CW.[CWD.OUTPUT]) OTE(MV_MV31R_D) ,XIC(S:FS) [OTU(MV_MV31R.CW.[CWD.MANUAL]) ,LEQ(MV_MV31R.CheckTime,0) MOV(Default_Check_Time,MV_MV31R.CheckTime) ] ,[[XIC(MV_MV31R_R) XIO(Item_Simulation_Flag) ,XIC(Item_Simulation_Flag) [XIC(MV_MV31R.CW.[CWD.OUTPUT]) XIO(MV_MV31R.CW.[CWD.SIMFAIL]) ,XIO(MV_MV31R.CW.[CWD.OUTPUT]) XIC(MV_MV31R.CW.[CWD.SIMFAIL]) ] ] OTE(MV_MV31R.CW.[CWD.RUNFB]) ,[XIC(Item_Simulation_Flag) ,XIC(MV_MV31R.CW.[CWD.CHECKOFF]) ,XIC(Unused_Healthy_Feedback) ] OTE(MV_MV31R.CW.[CWD.HEALTHYFB]) ,[XIC(Item_Simulation_Flag) ,XIC(MV_MV31R.CW.[CWD.CHECKOFF]) ,XIC(Unused_NotTripped_Feedback) ] OTE(MV_MV31R.CW.[CWD.NOTTRIPPEDFB]) ] ,[XIC(MV_MV31R.CW.[CWD.AUTODRV]) XIO(MV_MV31R.CW.[CWD.PREVSCAN]) ,XIO(MV_MV31R.CW.[CWD.AUTODRV]) XIC(MV_MV31R.CW.[CWD.PREVSCAN]) ] CLR(MV_MV31R.CheckTimer) ,XIC(One_Second_One_Scan) LES(MV_MV31R.CheckTimer,MV_MV31R.CheckTime) ADD(MV_MV31R.CheckTimer,1,MV_MV31R.CheckTimer) ,XIO(MV_MV31R.CW.[CWD.FAULT]) OTU(MV_MV31R.CW.[CWD.FAULTLOGGED]) ,[GEQ(MV_MV31R.CheckTimer,MV_MV31R.CheckTime) [XIC(MV_MV31R.CW.[CWD.OUTPUT]) XIO(MV_MV31R.CW.[CWD.RUNFB]) ,XIO(MV_MV31R.CW.[CWD.OUTPUT]) XIC(MV_MV31R.CW.[CWD.RUNFB]) ] ,XIO(MV_MV31R.CW.[CWD.HEALTHYFB]) ,XIO(MV_MV31R.CW.[CWD.NOTTRIPPEDFB]) ,XIC(MV_MV31R.CW.[CWD.FAULT]) XIC(Item_Faults_Are_Latched) ,XIC(MV_MV31R.CW.[CWD.HIGHLIGHT]) ] XIO(MV_MV31R.CW.[CWD.CHECKOFF]) XIO(Alarm_Reset) [OTE(MV_MV31R.CW.[CWD.FAULT]) ,ALMD(MV_MV31R_ALARM,0,0,0,0) ] ,XIC(MV_MV31R.CW.[CWD.OUTPUT]) OTE(MV_MV31R.CW.[CWD.PREVSCAN]) ,XIC(MV_MV31R.CW.[CWD.FAULT]) EQU(Scada_Pump_Fault_No,0) XIO(MV_MV31R.CW.[CWD.FAULTLOGGED]) [MOV(20001,Scada_Pump_Fault_No) ,OTL(MV_MV31R.CW.[CWD.FAULTLOGGED]) ] ,XIO(MV_MV31R.CW.[CWD.HEALTHYFB]) EQU(Scada_Pump_H_Fault_No,0) XIO(MV_MV31R.CW.[CWD.HEALTHYFAULTLOGGED]) [MOV(20001,Scada_Pump_H_Fault_No) ,OTL(MV_MV31R.CW.[CWD.HEALTHYFAULTLOGGED]) ] ,XIO(MV_MV31R.CW.[CWD.NOTTRIPPEDFB]) EQU(Scada_Pump_H_Fault_No,0) XIO(MV_MV31R.CW.[CWD.TRIPPEDFAULTLOGGED]) [MOV(20001,Scada_Pump_T_Fault_No) ,OTL(MV_MV31R.CW.[CWD.TRIPPEDFAULTLOGGED]) ] ];
   21: [NEQ(MV_MV32R.DriveBits,0) OTE(MV_MV32R.CW.[CWD.AUTODRV]) ,[XIC(MV_MV32R.CW.[CWD.AUTODRV]) XIO(MV_MV32R.CW.[CWD.MANUAL]) ,XIC(MV_MV32R.CW.[CWD.MANDRV]) XIC(MV_MV32R.CW.[CWD.MANUAL]) ] OTE(MV_MV32R.CW.[CWD.OUTPUT]) ,XIC(MV_MV32R.CW.[CWD.OUTPUT]) OTE(MV_MV32R_D) ,XIC(S:FS) [OTU(MV_MV32R.CW.[CWD.MANUAL]) ,LEQ(MV_MV32R.CheckTime,0) MOV(Default_Check_Time,MV_MV32R.CheckTime) ] ,[[XIC(MV_MV32R_R) XIO(Item_Simulation_Flag) ,XIC(Item_Simulation_Flag) [XIC(MV_MV32R.CW.[CWD.OUTPUT]) XIO(MV_MV32R.CW.[CWD.SIMFAIL]) ,XIO(MV_MV32R.CW.[CWD.OUTPUT]) XIC(MV_MV32R.CW.[CWD.SIMFAIL]) ] ] OTE(MV_MV32R.CW.[CWD.RUNFB]) ,[XIC(Item_Simulation_Flag) ,XIC(MV_MV32R.CW.[CWD.CHECKOFF]) ,XIC(Unused_Healthy_Feedback) ] OTE(MV_MV32R.CW.[CWD.HEALTHYFB]) ,[XIC(Item_Simulation_Flag) ,XIC(MV_MV32R.CW.[CWD.CHECKOFF]) ,XIC(Unused_NotTripped_Feedback) ] OTE(MV_MV32R.CW.[CWD.NOTTRIPPEDFB]) ] ,[XIC(MV_MV32R.CW.[CWD.AUTODRV]) XIO(MV_MV32R.CW.[CWD.PREVSCAN]) ,XIO(MV_MV32R.CW.[CWD.AUTODRV]) XIC(MV_MV32R.CW.[CWD.PREVSCAN]) ] CLR(MV_MV32R.CheckTimer) ,XIC(One_Second_One_Scan) LES(MV_MV32R.CheckTimer,MV_MV32R.CheckTime) ADD(MV_MV32R.CheckTimer,1,MV_MV32R.CheckTimer) ,XIO(MV_MV32R.CW.[CWD.FAULT]) OTU(MV_MV32R.CW.[CWD.FAULTLOGGED]) ,[GEQ(MV_MV32R.CheckTimer,MV_MV32R.CheckTime) [XIC(MV_MV32R.CW.[CWD.OUTPUT]) XIO(MV_MV32R.CW.[CWD.RUNFB]) ,XIO(MV_MV32R.CW.[CWD.OUTPUT]) XIC(MV_MV32R.CW.[CWD.RUNFB]) ] ,XIO(MV_MV32R.CW.[CWD.HEALTHYFB]) ,XIO(MV_MV32R.CW.[CWD.NOTTRIPPEDFB]) ,XIC(MV_MV32R.CW.[CWD.FAULT]) XIC(Item_Faults_Are_Latched) ,XIC(MV_MV32R.CW.[CWD.HIGHLIGHT]) ] XIO(MV_MV32R.CW.[CWD.CHECKOFF]) XIO(Alarm_Reset) [OTE(MV_MV32R.CW.[CWD.FAULT]) ,ALMD(MV_MV32R_ALARM,0,0,0,0) ] ,XIC(MV_MV32R.CW.[CWD.OUTPUT]) OTE(MV_MV32R.CW.[CWD.PREVSCAN]) ,XIC(MV_MV32R.CW.[CWD.FAULT]) EQU(Scada_Pump_Fault_No,0) XIO(MV_MV32R.CW.[CWD.FAULTLOGGED]) [MOV(20001,Scada_Pump_Fault_No) ,OTL(MV_MV32R.CW.[CWD.FAULTLOGGED]) ] ,XIO(MV_MV32R.CW.[CWD.HEALTHYFB]) EQU(Scada_Pump_H_Fault_No,0) XIO(MV_MV32R.CW.[CWD.HEALTHYFAULTLOGGED]) [MOV(20001,Scada_Pump_H_Fault_No) ,OTL(MV_MV32R.CW.[CWD.HEALTHYFAULTLOGGED]) ] ,XIO(MV_MV32R.CW.[CWD.NOTTRIPPEDFB]) EQU(Scada_Pump_H_Fault_No,0) XIO(MV_MV32R.CW.[CWD.TRIPPEDFAULTLOGGED]) [MOV(20001,Scada_Pump_T_Fault_No) ,OTL(MV_MV32R.CW.[CWD.TRIPPEDFAULTLOGGED]) ] ];
   22: [NEQ(MV_MV33R.DriveBits,0) OTE(MV_MV33R.CW.[CWD.AUTODRV]) ,[XIC(MV_MV33R.CW.[CWD.AUTODRV]) XIO(MV_MV33R.CW.[CWD.MANUAL]) ,XIC(MV_MV33R.CW.[CWD.MANDRV]) XIC(MV_MV33R.CW.[CWD.MANUAL]) ] OTE(MV_MV33R.CW.[CWD.OUTPUT]) ,XIC(MV_MV33R.CW.[CWD.OUTPUT]) OTE(MV_MV33R_D) ,XIC(S:FS) [OTU(MV_MV33R.CW.[CWD.MANUAL]) ,LEQ(MV_MV33R.CheckTime,0) MOV(Default_Check_Time,MV_MV33R.CheckTime) ] ,[[XIC(MV_MV33R_R) XIO(Item_Simulation_Flag) ,XIC(Item_Simulation_Flag) [XIC(MV_MV33R.CW.[CWD.OUTPUT]) XIO(MV_MV33R.CW.[CWD.SIMFAIL]) ,XIO(MV_MV33R.CW.[CWD.OUTPUT]) XIC(MV_MV33R.CW.[CWD.SIMFAIL]) ] ] OTE(MV_MV33R.CW.[CWD.RUNFB]) ,[XIC(Item_Simulation_Flag) ,XIC(MV_MV33R.CW.[CWD.CHECKOFF]) ,XIC(Unused_Healthy_Feedback) ] OTE(MV_MV33R.CW.[CWD.HEALTHYFB]) ,[XIC(Item_Simulation_Flag) ,XIC(MV_MV33R.CW.[CWD.CHECKOFF]) ,XIC(Unused_NotTripped_Feedback) ] OTE(MV_MV33R.CW.[CWD.NOTTRIPPEDFB]) ] ,[XIC(MV_MV33R.CW.[CWD.AUTODRV]) XIO(MV_MV33R.CW.[CWD.PREVSCAN]) ,XIO(MV_MV33R.CW.[CWD.AUTODRV]) XIC(MV_MV33R.CW.[CWD.PREVSCAN]) ] CLR(MV_MV33R.CheckTimer) ,XIC(One_Second_One_Scan) LES(MV_MV33R.CheckTimer,MV_MV33R.CheckTime) ADD(MV_MV33R.CheckTimer,1,MV_MV33R.CheckTimer) ,XIO(MV_MV33R.CW.[CWD.FAULT]) OTU(MV_MV33R.CW.[CWD.FAULTLOGGED]) ,[GEQ(MV_MV33R.CheckTimer,MV_MV33R.CheckTime) [XIC(MV_MV33R.CW.[CWD.OUTPUT]) XIO(MV_MV33R.CW.[CWD.RUNFB]) ,XIO(MV_MV33R.CW.[CWD.OUTPUT]) XIC(MV_MV33R.CW.[CWD.RUNFB]) ] ,XIO(MV_MV33R.CW.[CWD.HEALTHYFB]) ,XIO(MV_MV33R.CW.[CWD.NOTTRIPPEDFB]) ,XIC(MV_MV33R.CW.[CWD.FAULT]) XIC(Item_Faults_Are_Latched) ,XIC(MV_MV33R.CW.[CWD.HIGHLIGHT]) ] XIO(MV_MV33R.CW.[CWD.CHECKOFF]) XIO(Alarm_Reset) [OTE(MV_MV33R.CW.[CWD.FAULT]) ,ALMD(MV_MV33R_ALARM,0,0,0,0) ] ,XIC(MV_MV33R.CW.[CWD.OUTPUT]) OTE(MV_MV33R.CW.[CWD.PREVSCAN]) ,XIC(MV_MV33R.CW.[CWD.FAULT]) EQU(Scada_Pump_Fault_No,0) XIO(MV_MV33R.CW.[CWD.FAULTLOGGED]) [MOV(20001,Scada_Pump_Fault_No) ,OTL(MV_MV33R.CW.[CWD.FAULTLOGGED]) ] ,XIO(MV_MV33R.CW.[CWD.HEALTHYFB]) EQU(Scada_Pump_H_Fault_No,0) XIO(MV_MV33R.CW.[CWD.HEALTHYFAULTLOGGED]) [MOV(20001,Scada_Pump_H_Fault_No) ,OTL(MV_MV33R.CW.[CWD.HEALTHYFAULTLOGGED]) ] ,XIO(MV_MV33R.CW.[CWD.NOTTRIPPEDFB]) EQU(Scada_Pump_H_Fault_No,0) XIO(MV_MV33R.CW.[CWD.TRIPPEDFAULTLOGGED]) [MOV(20001,Scada_Pump_T_Fault_No) ,OTL(MV_MV33R.CW.[CWD.TRIPPEDFAULTLOGGED]) ] ];
   23: [NEQ(MV_MV34R.DriveBits,0) OTE(MV_MV34R.CW.[CWD.AUTODRV]) ,[XIC(MV_MV34R.CW.[CWD.AUTODRV]) XIO(MV_MV34R.CW.[CWD.MANUAL]) ,XIC(MV_MV34R.CW.[CWD.MANDRV]) XIC(MV_MV34R.CW.[CWD.MANUAL]) ] OTE(MV_MV34R.CW.[CWD.OUTPUT]) ,XIC(MV_MV34R.CW.[CWD.OUTPUT]) OTE(MV_MV34R_D) ,XIC(S:FS) [OTU(MV_MV34R.CW.[CWD.MANUAL]) ,LEQ(MV_MV34R.CheckTime,0) MOV(Default_Check_Time,MV_MV34R.CheckTime) ] ,[[XIC(MV_MV34R_R) XIO(Item_Simulation_Flag) ,XIC(Item_Simulation_Flag) [XIC(MV_MV34R.CW.[CWD.OUTPUT]) XIO(MV_MV34R.CW.[CWD.SIMFAIL]) ,XIO(MV_MV34R.CW.[CWD.OUTPUT]) XIC(MV_MV34R.CW.[CWD.SIMFAIL]) ] ] OTE(MV_MV34R.CW.[CWD.RUNFB]) ,[XIC(Item_Simulation_Flag) ,XIC(MV_MV34R.CW.[CWD.CHECKOFF]) ,XIC(Unused_Healthy_Feedback) ] OTE(MV_MV34R.CW.[CWD.HEALTHYFB]) ,[XIC(Item_Simulation_Flag) ,XIC(MV_MV34R.CW.[CWD.CHECKOFF]) ,XIC(Unused_NotTripped_Feedback) ] OTE(MV_MV34R.CW.[CWD.NOTTRIPPEDFB]) ] ,[XIC(MV_MV34R.CW.[CWD.AUTODRV]) XIO(MV_MV34R.CW.[CWD.PREVSCAN]) ,XIO(MV_MV34R.CW.[CWD.AUTODRV]) XIC(MV_MV34R.CW.[CWD.PREVSCAN]) ] CLR(MV_MV34R.CheckTimer) ,XIC(One_Second_One_Scan) LES(MV_MV34R.CheckTimer,MV_MV34R.CheckTime) ADD(MV_MV34R.CheckTimer,1,MV_MV34R.CheckTimer) ,XIO(MV_MV34R.CW.[CWD.FAULT]) OTU(MV_MV34R.CW.[CWD.FAULTLOGGED]) ,[GEQ(MV_MV34R.CheckTimer,MV_MV34R.CheckTime) [XIC(MV_MV34R.CW.[CWD.OUTPUT]) XIO(MV_MV34R.CW.[CWD.RUNFB]) ,XIO(MV_MV34R.CW.[CWD.OUTPUT]) XIC(MV_MV34R.CW.[CWD.RUNFB]) ] ,XIO(MV_MV34R.CW.[CWD.HEALTHYFB]) ,XIO(MV_MV34R.CW.[CWD.NOTTRIPPEDFB]) ,XIC(MV_MV34R.CW.[CWD.FAULT]) XIC(Item_Faults_Are_Latched) ,XIC(MV_MV34R.CW.[CWD.HIGHLIGHT]) ] XIO(MV_MV34R.CW.[CWD.CHECKOFF]) XIO(Alarm_Reset) [OTE(MV_MV34R.CW.[CWD.FAULT]) ,ALMD(MV_MV34R_ALARM,0,0,0,0) ] ,XIC(MV_MV34R.CW.[CWD.OUTPUT]) OTE(MV_MV34R.CW.[CWD.PREVSCAN]) ,XIC(MV_MV34R.CW.[CWD.FAULT]) EQU(Scada_Pump_Fault_No,0) XIO(MV_MV34R.CW.[CWD.FAULTLOGGED]) [MOV(20001,Scada_Pump_Fault_No) ,OTL(MV_MV34R.CW.[CWD.FAULTLOGGED]) ] ,XIO(MV_MV34R.CW.[CWD.HEALTHYFB]) EQU(Scada_Pump_H_Fault_No,0) XIO(MV_MV34R.CW.[CWD.HEALTHYFAULTLOGGED]) [MOV(20001,Scada_Pump_H_Fault_No) ,OTL(MV_MV34R.CW.[CWD.HEALTHYFAULTLOGGED]) ] ,XIO(MV_MV34R.CW.[CWD.NOTTRIPPEDFB]) EQU(Scada_Pump_H_Fault_No,0) XIO(MV_MV34R.CW.[CWD.TRIPPEDFAULTLOGGED]) [MOV(20001,Scada_Pump_T_Fault_No) ,OTL(MV_MV34R.CW.[CWD.TRIPPEDFAULTLOGGED]) ] ];
